               IF (#TMP_dNextTail + 1) >= "DMAXGLASSDATASECTORS" THEN
                   #TMP_dNextTail := 0;
               ELSE
                   #TMP_dNextTail += 1;
               END_IF;

               #TMP_dValue_cmm := #INO_tRibbon.rgtGlassData[#TMP_dSourceIndex].rgtBuffer[#TMP_dNextTail].dEncoderValue_cmm - #INO_tEncoder.dActualEncoderCounter_cmm;

               IF (#TMP_dValue_cmm <= #INO_tRibbon.rgtGlassDataRequest[#TMP_dIndex].IN_dDistanceSnaproll_cmm) THEN

                   #INO_tRibbon.rgtGlassDataRequest[#TMP_dIndex].OUT_dGrossWidth_cmm := #INO_tRibbon.rgtGlassData[#TMP_dSourceIndex].rgtBuffer[#TMP_dNextTail].dGrossWidth_cmm;
                   #INO_tRibbon.rgtGlassDataRequest[#TMP_dIndex].OUT_dNetWidth_cmm := #INO_tRibbon.rgtGlassData[#TMP_dSourceIndex].rgtBuffer[#TMP_dNextTail].dNetWidth_cmm;
                   #INO_tRibbon.rgtGlassDataRequest[#TMP_dIndex].OUT_dGrossWander_cmm := #INO_tRibbon.rgtGlassData[#TMP_dSourceIndex].rgtBuffer[#TMP_dNextTail].dGrossWander_cmm;
                   #INO_tRibbon.rgtGlassDataRequest[#TMP_dIndex].OUT_dNetWander_cmm := #INO_tRibbon.rgtGlassData[#TMP_dSourceIndex].rgtBuffer[#TMP_dNextTail].dNetWander_cmm;

               ELSE
                   EXIT;
               END_IF;

           END_WHILE;
           //Setup data ready
           #INO_tRibbon.rgtGlassDataRequest[#TMP_dIndex].OUT_xDataReady := TRUE;
       END_IF;
   END_FOR;
END_REGION

REGION Network 8 (SCL): Evaluate glass break request
   FOR #TMP_dIndex := 0 TO "DMAXGLASSBREAKREQUEST_IND" DO

       #TMP_xGlassBreak := FALSE;

       IF #INO_tRibbon.rgtGlassBreakRequest[#TMP_dIndex].IN_xRequestGlassBreak AND NOT #INO_tRibbon.rgtGlassBreakRequest[#TMP_dIndex].OUT_xDataReady THEN

           //Evaluate the glass break machine, only the machine before the requested position 
           FOR #TMP_dBreakMachIndex := 0 TO #INO_tRibbon.dActualNumberGlassBreakMachine - 1 DO

               IF (#INO_tRibbon.rgtGlassBreakRequest[#TMP_dIndex].IN_dDistanceSnaproll_cmm >= #INO_tRibbon.rgtGlassBreak[#TMP_dBreakMachIndex].dDistSnapRoll_cmm) THEN
                   CONTINUE;
               END_IF;

               #TMP_xGlassBreak := #INO_tRibbon.rgtGlassBreak[#TMP_dBreakMachIndex].tLastDataBuffer.xGlassBreak;

               #TMP_dNextTail := #INO_tRibbon.rgtGlassBreak[#TMP_dBreakMachIndex].dBufferTail;

               WHILE (#TMP_dNextTail <> #INO_tRibbon.rgtGlassBreak[#TMP_dBreakMachIndex].dBufferHead)
                   AND (#INO_tRibbon.rgtGlassBreak[#TMP_dBreakMachIndex].dBufferHead <> -1) DO

                   IF (#TMP_dNextTail + 1) >= "DMAXGLASSBREAKSECTORS" THEN
                       #TMP_dNextTail := 0;
                   ELSE
                       #TMP_dNextTail += 1;
                   END_IF;

                   #TMP_dValue_cmm := #INO_tRibbon.rgtGlassBreak[#TMP_dBreakMachIndex].rgtBuffer[#TMP_dNextTail].dEncoderValue_cmm - #INO_tEncoder.dActualEncoderCounter_cmm;

                   IF (#TMP_dValue_cmm <= #INO_tRibbon.rgtGlassBreakRequest[#TMP_dIndex].IN_dDistanceSnaproll_cmm) THEN

                       //If the distance is less the snaproll, but greather the safety band. In case of glass break the system will not overwrite the information
                       IF (#TMP_dValue_cmm < #INO_tRibbon.rgtGlassBreakRequest[#TMP_dIndex].IN_dDistanceSnaproll_cmm - #INO_tRibbon.rgtGlassBreakRequest[#TMP_dIndex].IN_dDownstreamOffset_cmm) THEN
                           #TMP_xGlassBreak := #INO_tRibbon.rgtGlassBreak[#TMP_dBreakMachIndex].rgtBuffer[#TMP_dNextTail].xGlassBreak;
                       ELSE
                           IF NOT #TMP_xGlassBreak THEN
                               #TMP_xGlassBreak := #INO_tRibbon.rgtGlassBreak[#TMP_dBreakMachIndex].rgtBuffer[#TMP_dNextTail].xGlassBreak;
                           END_IF;
                       END_IF;

                   ELSE

                       //The position is greather, but still on the position window
                       IF (#TMP_dValue_cmm <= #INO_tRibbon.rgtGlassBreakRequest[#TMP_dIndex].IN_dDistanceSnaproll_cmm + #INO_tRibbon.rgtGlassBreakRequest[#TMP_dIndex].IN_dUpstreamOffset_cmm) THEN
                           IF NOT #TMP_xGlassBreak THEN
                               #TMP_xGlassBreak := #INO_tRibbon.rgtGlassBreak[#TMP_dBreakMachIndex].rgtBuffer[#TMP_dNextTail].xGlassBreak;
                           END_IF;
                       ELSE
                           EXIT; //Exit the while
                       END_IF;

                   END_IF;

               END_WHILE;

               IF #TMP_xGlassBreak THEN
                   EXIT;
               END_IF;
           END_FOR;

           #INO_tRibbon.rgtGlassBreakRequest[#TMP_dIndex].OUT_xDataReady := TRUE;
           #INO_tRibbon.rgtGlassBreakRequest[#TMP_dIndex].OUT_xGlassBreak := #TMP_xGlassBreak;

       END_IF;
   END_FOR;
END_REGION
END_FUNCTION_BLOCK

// folder: 03_Programs_Logics/MCC1200/18_ISRA

FUNCTION_BLOCK "FB_ISRA5D"   // FB21, LAD
{ S7_Optimized_Access := 'TRUE' }
VERSION : 0.1
   VAR_INPUT
      IN_xCycleON : Bool;   // Cycle ON
      IN_xCycleONDel : Bool;   // Delayed cycle ON signal
      IN_dGlassBreakIndexGet : DInt;   // Glass break index get
      IN_xGeneralReset : Bool;   // General reset
      IN_xResetAlarms : Bool;   // Reset alarms
      IN_xFaultsEnabled : Bool;   // Faults enabled
      IN_tInterfaceID : Hw_Any;   // Interface ID
      IN_tID : Conn_Ouc;   // Connection ID
      IN_uiLocalPort : UInt;   // Local port
      IN_dGlassDataMachineIndex : DInt;   // Glass data machine index
      IN_dGlassDataUpdateMachineIndex : DInt;   // Glass data update machine index
      IN_xSimulationActive : Bool;   // Enable simulation (EXPERT USER)
      IN_xScannerON : Bool;
   END_VAR
   VAR_OUTPUT
      OUT_xGlassBreak : Bool;
   END_VAR
   VAR_IN_OUT
      INO_tFBAddDefect : "FB_Defects_Add_V1.00";   // Add defect on buffer
      INO_xDefectBufferFull : Bool;   // Defect buffer full
      INO_tEncoder : "UDT_Encoder";   // Encoder data
      INO_tRibbon : "UDT_RibbonData";   // Ribbon data
      INO_tOptManager : "FB_OptManager_V1.00";   // Optimizer manager
      INO_tCaps : "UDT_CapData_Tracking";   // Caps data
      INO_OB_Init : "GP_OB_Initialize";
   END_VAR
   VAR
      tALM : Struct   // HMI Alarms
         tS : Struct   // Stopping faults
            xNotSyncro : Bool;   // Machine not syncronized {X|X|X|X|O}
            xScannerNotConnected : Bool;   // Scanner not connected {X|X|X|X|O}
            xSpare_2 : Bool;
            xSpare_3 : Bool;
            xSpare_4 : Bool;
            xSpare_5 : Bool;
            xSpare_6 : Bool;
            xSpare_7 : Bool;
            xSpare_8 : Bool;
            xSpare_9 : Bool;
            xSpare_10 : Bool;
            xSpare_11 : Bool;
            xSpare_12 : Bool;
            xSpare_13 : Bool;
            xSpare_14 : Bool;
            xSpare_15 : Bool;
            xSpare_16 : Bool;
            xSpare_17 : Bool;
            xSpare_18 : Bool;
            xSpare_19 : Bool;
            xSpare_20 : Bool;
            xSpare_21 : Bool;
            xSpare_22 : Bool;
            xSpare_23 : Bool;
            xSpare_24 : Bool;
            xSpare_25 : Bool;
            xSpare_26 : Bool;
            xSpare_27 : Bool;
            xSpare_28 : Bool;
            xSpare_29 : Bool;
            xSpare_30 : Bool;
            xSpare_31 : Bool;
         END_STRUCT;
         tF : Struct   // Faults
            xUTelMissing : Bool;   // U telegram missing {X|X|X|X|O}
            xSTelMissing : Bool;   // S telegram missing {X|X|X|X|O}
            xCTelMissing : Bool;   // C telegram missing {X|X|X|X|O}
            xYTelMissing : Bool;   // Y telegram missing {X|X|X|X|O}
            xBTelMissing : Bool;   // B telegram missing {X|X|X|X|O}
            xSpare_5 : Bool;
            xSpare_6 : Bool;
            xSpare_7 : Bool;
            xSpare_8 : Bool;
            xSpare_9 : Bool;
            xSpare_10 : Bool;
            xSpare_11 : Bool;
            xSpare_12 : Bool;
            xSpare_13 : Bool;
            xSpare_14 : Bool;
            xSpare_15 : Bool;
            xSpare_16 : Bool;
            xSpare_17 : Bool;
            xSpare_18 : Bool;
            xSpare_19 : Bool;
            xSpare_20 : Bool;
            xSpare_21 : Bool;
            xSpare_22 : Bool;
            xSpare_23 : Bool;
            xSpare_24 : Bool;
            xSpare_25 : Bool;
            xSpare_26 : Bool;
            xSpare_27 : Bool;
            xSpare_28 : Bool;
            xSpare_29 : Bool;
            xSpare_30 : Bool;
            xSpare_31 : Bool;
         END_STRUCT;
         tW : Struct   // Warnings
            xSpare_0 : Bool;
            xSpare_1 : Bool;
            xSpare_2 : Bool;
            xSpare_3 : Bool;
            xSpare_4 : Bool;
            xSpare_5 : Bool;
            xSpare_6 : Bool;
            xSpare_7 : Bool;
            xSpare_8 : Bool;
            xSpare_9 : Bool;
            xSpare_10 : Bool;
            xSpare_11 : Bool;
            xSpare_12 : Bool;
            xSpare_13 : Bool;
            xSpare_14 : Bool;
            xSpare_15 : Bool;
            xSpare_16 : Bool;
            xSpare_17 : Bool;
            xSpare_18 : Bool;
            xSpare_19 : Bool;
            xSpare_20 : Bool;
            xSpare_21 : Bool;
            xSpare_22 : Bool;
            xSpare_23 : Bool;
            xSpare_24 : Bool;
            xSpare_25 : Bool;
            xSpare_26 : Bool;
            xSpare_27 : Bool;
            xSpare_28 : Bool;
            xSpare_29 : Bool;
            xSpare_30 : Bool;
            xSpare_31 : Bool;
         END_STRUCT;
      END_STRUCT;
   END_VAR
   VAR RETAIN
      tHMR : Struct
         dInspectionStatus : DInt;   // Inspection status (1=Disabled 3=Enabled 4=Wait first syncro 7=Anomaly ) {X|X|X|X|O}
         xScannerON : Bool;   // xScannerON {X|X|X|X|O}
         dDistSnapRoll_cmm : DInt;   // Distance from snaproll [mm/100] {mm/100|mm|X|X|O}
         dDistCenterLine_cmm : DInt;   // Distance from center line [mm/100] {mm/100|mm|X|X|O}
         dCurrentGrossWidth_cmm : DInt;   // Gross width [mm/100] {mm/100|mm|X|X|O}
         dCurrentNetWidth_cmm : DInt;   // Net width [mm/100] {mm/100|mm|X|X|O}
         dCurrentGrossWander_cmm : DInt;   // Gross wander [mm/100] {mm/100|mm|X|X|O}
         dCurrentNetWander_cmm : DInt;   // Net wander [mm/100] {mm/100|mm|X|X|O}
      END_STRUCT;
      tHMW : Struct   // HMI Write
         xAutoInspEnabled : Bool;   // Automatic inspection enabled {X|X|X|X|O}
         xUpdDistSnaproll : Bool;   // Update distance from snaproll {X|X|X|X|O}
         xUpdDistCenterLine : Bool;   // Update distance from center line {X|X|X|X|O}
         xCalibPosition : Bool;   // Calibrate defect position {X|X|X|X|O}
         dCalibDefRealXPos_cmm : DInt;   // Calibration defect real X position [mm/100] {mm/100|mm|0|7000|O}
         dCalibDefRealYPos_cmm : DInt;   // Calibration defect real Y position [mm/100] {mm/100|mm|0|4000|O}
         dCalibDefTeoXPos_cmm : DInt;   // Calibration defect theorical X position [mm/100] {mm/100|mm|0|7000|O}
         dCalibDefTeoYPos_cmm : DInt;   // Calibration defect theorical Y position [mm/100] {mm/100|mm|0|4000|O}
         dDistSnapRoll_cmm : DInt;   // Distance from snaproll [mm/100] {mm/100|mm|0|70000|O}
         dDistCenterLine_cmm : DInt;   // Distance from center line [mm/100] {mm/100|mm|-4000|4000|O}
      END_STRUCT;
   END_VAR
   VAR
      tPhNet : Struct   // Network phases
         xSendInProgress : Bool;   // Send data in progress
         xEndSendInProgress : Bool;   // End send data in progress
         xSpare_2 : Bool;
         xSpare_3 : Bool;
         xSpare_4 : Bool;
         xSpare_5 : Bool;
         xSpare_6 : Bool;
         xSpare_7 : Bool;
         xSpare_8 : Bool;
         xSpare_9 : Bool;
         xSpare_10 : Bool;
         xSpare_11 : Bool;
         xSpare_12 : Bool;
         xSpare_13 : Bool;
         xSpare_14 : Bool;
         xSpare_15 : Bool;
         xSpare_16 : Bool;
         xSpare_17 : Bool;
         xSpare_18 : Bool;
         xSpare_19 : Bool;
         xSpare_20 : Bool;
         xSpare_21 : Bool;
         xSpare_22 : Bool;
         xSpare_23 : Bool;
         xSpare_24 : Bool;
         xSpare_25 : Bool;
         xSpare_26 : Bool;
         xSpare_27 : Bool;
         xSpare_28 : Bool;
         xSpare_29 : Bool;
         xSpare_30 : Bool;
         xSpare_31 : Bool;
      END_STRUCT;
      tPh : Struct   // Machine phases
         xWaitSyncroData : Bool;   // Wait syncro data
         xEndWaitSyncroData : Bool;   // End wait syncro data
         xSpare_2 : Bool;
         xSpare_3 : Bool;
         xSpare_4 : Bool;
         xSpare_5 : Bool;
         xSpare_6 : Bool;
         xSpare_7 : Bool;
         xSpare_8 : Bool;
         xSpare_9 : Bool;
         xSpare_10 : Bool;
         xSpare_11 : Bool;
         xSpare_12 : Bool;
         xSpare_13 : Bool;
         xSpare_14 : Bool;
         xSpare_15 : Bool;
         xSpare_16 : Bool;
         xSpare_17 : Bool;
         xSpare_18 : Bool;
         xSpare_19 : Bool;
         xSpare_20 : Bool;
         xSpare_21 : Bool;
         xSpare_22 : Bool;
         xSpare_23 : Bool;
         xSpare_24 : Bool;
         xSpare_25 : Bool;
         xSpare_26 : Bool;
         xSpare_27 : Bool;
         xSpare_28 : Bool;
         xSpare_29 : Bool;
         xSpare_30 : Bool;
         xSpare_31 : Bool;
      END_STRUCT;
      ST_xMachineSyncronized : Bool;   // Machine is syncronized
      ST_xStoppedFaults : Bool;   // Stopped faults
      ST_xFaults : Bool;   // Faults
      ST_xWarning : Bool;   // Warnings
      ST_xGlassBreak : Bool;   // Glass break
      OS_xSyncroOutLimits : Bool;   // OS.Syncro outside limits
      OS_xSyncroTimeout : Bool;   // OS.Syncro timeout
      AUX_xTelegramError : Bool;   // Telegram error
      AUX_xTelegramYError : Bool;   // Telegram Y error
      AUX_xTelegramBError : Bool;   // Telegram B error
      AUX_xTelegramCError : Bool;   // Telegram C error
      AUX_xTelegramSError : Bool;   // Telegram S error
      AUX_xTelegramUError : Bool;   // Telegram U error
      AUX_xTelegramYMissing : Bool;   // Telegram Y missing
      AUX_xTelegramBMissing : Bool;   // Telegram B missing
      AUX_xTelegramCMissing : Bool;   // Telegram C missing
      AUX_xTelegramSMissing : Bool;   // Telegram S missing
      AUX_xTelegramUMissing : Bool;   // Telegram U missing
      AUX_tUTelegram : Struct   // U telegram
         dTelCounter : DInt;   // Telegram counter [0..65535]
         dFeedPulse_mm : DInt;   // Feeding pulse counter [mm]
         dDefPos_mm : DInt;   // Defect position [mm]
         dDefLengthTot_um : DInt;   // Defect length total [um]
         dDefWidthTot_um : DInt;   // Defect width total [um]
         dDefLengthCore_um : DInt;   // Defect length core [um]
         dDefWidthCore_um : DInt;   // Defect width core [um]
         dDefLengthDef_um : DInt;   // Defect length deformation [um]
         dDefWidthDef_um : DInt;   // Defect width deformation [um]
         dClass : DInt;   // Defect class [01..99]
         dType : DInt;   // Defect type [01..99]
         dPLCPosCount_cmm : DInt;   // PLC Position counter [mm/100]
         dPLCYPos_cmm : DInt;   // PLC Y position value [mm/100]
         strDefectID : String;   // Defect ID string
      END_STRUCT;
      AUX_tYTelegram : Struct   // Y telegram
         dTelCounter : DInt;   // Telegram counter [0..65535]
         dFeedPulse_mm : DInt;   // Feeding pulse counter [mm]
         dInLimit_mm : DInt;   // Inner limit of the observation area [mm]
         dOutLimit_mm : DInt;   // Outer limit o fthe observation area [mm]
         dInLimitUsable_mm : DInt;   // Inner limit of the usable glass width [mm]
         dOutLimitUsable_mm : DInt;   // Outer limit of the usable glass width [mm]
         dInLimitGross_mm : DInt;   // Inner gross glass width [mm]
         dOutLimitGross_mm : DInt;   // Outer gross glass width [mm]
         dCenterOrientInTop_mm : DInt;   // Center orientated position of the inner toproller [mm]
         dEdgeOrientInTop_mm : DInt;   // Edge orientated position of the inner toproller [mm]
         dCenterOrientOutTop_mm : DInt;   // Center orientated position of the outer toproller [mm]
         dEdgeOrientOutTop_mm : DInt;   // Edge orientated position of the outer toproll [mm]
         dPLCPosCount_cmm : DInt;   // PLC Position counter [mm/100]
         dPLCYPos_cmm : DInt;   // PLC Y position value [mm/100]
      END_STRUCT;
      AUX_tCTelegram : Struct   // C Telegram
         dTelCounter : DInt;   // Telegram counter [0..65535]
         dFeedPulseStart_mm : DInt;   // Feeding pulse start counter [mm]
         dFeedPulseEnd_mm : DInt;   // Feeding pulse end counter [mm]
         dBeginAreaY_mm : DInt;   // Begin area Y [mm]
         dEndAreaY_mm : DInt;   // End area Y [mm]
         dPLCPosCountStart_cmm : DInt;   // PLC Position counter start [mm/100]
         dPLCPosCountEnd_cmm : DInt;   // PLC Position counter end [mm/100]
         dPLCYPosStart_cmm : DInt;   // PLC Y position value start [mm/100]
         dPLCYPosEnd_cmm : DInt;   // PLC Y position value end [mm/100]
         dPLCClusterLength_um : DInt;   // PLC Cluster length [um]
         dPLCClusterWidth_um : DInt;   // PLC Cluster width [um]
      END_STRUCT;
      AUX_tBTelegram : Struct   // B Telegram
         dTelCounter : DInt;   // Telegram counter [0..65535]
         dFeedPulse_mm : DInt;   // Feeding pulse counter [mm]
         xNewTelegram : Bool;   // New telegram received
      END_STRUCT;
      AUX_tSTelegram : Struct   // S Telegram
         dTelCounter : DInt;   // Telegram counter [0..65535]
         dFeedPulse_mm : DInt;   // Feeding pulse counter [mm]
         xNewTelegram : Bool;   // New telegram received
      END_STRUCT;
      AUX_tWTelegram : Struct   // T Telegram
         dTelCounter : DInt;   // Telegram counter [0..65535]
         dFeedPulse_mm : DInt;   // Feeding pulse counter [mm]
         dGrossWidthMin_mm : DInt;   // Gross width min [mm]
         dGrossWidthMax_mm : DInt;   // Gross width max [mm]
         dCutToolOpSide_mm : DInt;   // Cut tool opside [mm]
         dCutToolOppoOpSide_mm : DInt;   // Cut tool opposite operator side [mm]
         xNewTelegram : Bool;   // New telegram received
      END_STRUCT;
      AUX_dISRAValidCountMeter_mm : DInt;   // Last valid isra counter on meter [mm]
      AUX_dPLCValidCountMeter_cmm : DInt;   // Last valid PLC counter on meter [mm/100]
      AUX_rgcReceiveBuffer : Array[0..#DRECV_BUFFER_MAX_IND] of Char;   // Receive buffer
      AUX_dNumCharRecvBuffer : DInt;   // Number of char on the receive buffer
      AUX_rgsWTelegram : Array[0..#DNUMCHAR_TEL_W_INDEX] of Char;   // T Telegram char array
      AUX_tConnData : TCON_IP_v4;   // Connection data structure
      FB_TSend : TSEND_C;   // FB send
      FB_TRecv : TRCV_C;   // FB receive
      AUX_xResetSendConnection : Bool;   // Reset send connection
      AUX_rgcReceiveTempBuffer : Array[0..#DRECV_BUFFER_TEMP_IND] of Char;   // Temporary receive buffer
      tmON_SendTimeout : "UDT_IECTON_V1.00";   // Send timeout
      AUX_xSimDecModeGWidth : Bool;   // SIMULATION - Decrement mode gross width
      AUX_xSimIncModeGWidth : Bool;   // SIMULATION - Increment mode gross width
      AUX_xSimDecModeNWidth : Bool;   // SIMULATION - Decrement mode net width
      AUX_xSimIncModeNWidth : Bool;   // SIMULATION - Decrement mode net width
      AUX_xSimDecModeWander : Bool;   // SIMULATION - Decrement mode wander
      AUX_xSimIncModeWander : Bool;   // SIMULATION - Decrement mode wander
   END_VAR
   VAR RETAIN
      AUX_dSimGrossWidth_cmm : DInt;   // SIMULATION - Gross width [mm/100]
      AUX_dSimNetWidth_cmm : DInt;   // SIMULATION - Net width [mm/100]
      AUX_dSimWander_cmm : DInt;   // SIMULATION - Wander [mm/100]
   END_VAR
   VAR_TEMP
      TMP_dwValue : DWord;
      TMP_dIndex : DInt;
      TMP_dCharCounter : DInt;
      TMP_dTelCount : DInt;
      TMP_strValue : String;
      TMP_dCountPos_cmm : DInt;
      TMP_iRetVal : Int;
      TMP_dValue_cmm : DInt;
      TMP_xDummy : Bool;
      TMP_iStrLength : Int;
      TMP_uiMovedChar : UInt;
      TMP_xEnableReceive : Bool;
   END_VAR
   VAR CONSTANT
      DRECV_BUFFER_MAX : DInt := 5000;   // Maximum number of character on the receive buffer
      DRECV_BUFFER_MAX_IND : DInt := 4999;   // Maximum number of character on the receive buffer index
      DRECV_BUFFER_TEMP : DInt := 1000;   // Maximum number of character on the temporary receive buffer
      DRECV_BUFFER_TEMP_IND : DInt := 999;   // Maximum number of character on the temporary receive buffer index
      STR_CR : Char := '$R';   // CR
      STR_LF : Char := '$L';   // LF
      DNUMCHAR_TEL_U : DInt := 106;   // Number of char U telegram
      DNUMCHAR_TEL_C : DInt := 36;   // Number of char C telegram
      DNUMCHAR_TEL_Y : DInt := 75;   // Number of char Y telegram
      DNUMCHAR_TEL_B_S : DInt := 15;   // Number of char B - S telegram
      DCLUSTER_CLASS : DInt := 21;   // Cluster defect used class
      DCLUSTER_SUBTYPE : DInt := 1004;   // Cluster defect subtype
      DNUMCHAR_TEL_W : DInt := 39;   // Number of char W telegram
      DNUMCHAR_TEL_W_INDEX : DInt := 38;   // Number of char W telegram index
      DISRADEADPOINT_CMM : DInt := 250000;   // ISRA Dead point position quota [mm/100]
      CONST_DBREAKDOWNOFF_CMM : DInt := 100000;   // Break downstream offset [mm/100]
      CONST_DBREAKUPOFF_CMM : DInt := 100000;   // Break upstream offset [mm/100]
      BCONNTYPE : Byte := 16#0B;   // Optimizer connection type
      DSIM_MINGROSSWIDTH_CMM : DInt := 340000;   // Simulation minimum gross width [mm/100]
      DSIM_MAXGROSSWIDTH_CMM : DInt := 350000;   // Simulation maximum gross width [mm/100]
      DSIM_MINNETWIDTH_CMM : DInt := 330000;   // Simulation minimum net width [mm/100]
      DSIM_MAXNETWIDTH_CMM : DInt := 340000;   // Simulation maximum net width [mm/100]
      DSIM_MINNETWANDER_CMM : DInt := -20000;   // Simulation minimum net wander [mm/100]
      DSIM_MAXNETWANDER_CMM : DInt := 20000;   // Simulation maximum net wander [mm/100]
   END_VAR
   VAR_TEMP   // added for the SCL form of the ladder/FBD networks
      _w1 : Bool;
   END_VAR
BEGIN

REGION Network 1: ####_CONSTANTS_####
END_REGION

REGION Network 2 (SCL): General reset actions
   IF #IN_xGeneralReset THEN

       #AUX_tConnData.InterfaceId := #IN_tInterfaceID;
       #AUX_tConnData.ID := #IN_tID;
       #AUX_tConnData.ConnectionType := #BCONNTYPE;
       #AUX_tConnData.ActiveEstablished := FALSE;
       #AUX_tConnData.RemotePort := 0;
       #AUX_tConnData.LocalPort := #IN_uiLocalPort;

       #tPh.xWaitSyncroData := FALSE;
       #tPh.xEndWaitSyncroData := FALSE;

       #tPhNet.xSendInProgress := FALSE;
       #tPhNet.xEndSendInProgress := FALSE;

   END_IF;
END_REGION

REGION Network 3: ### ETHERNET RECEIVE DATA ###
END_REGION

REGION Network 4 (SCL): Manage send and receive
   #AUX_xResetSendConnection := #IN_xGeneralReset OR (#FB_TSend.s_TDIAG_Status.State <> b#16#04 AND #IN_xResetAlarms);

   #FB_TSend(REQ:=#tPhNet.xSendInProgress,
             CONT:=TRUE,
             LEN:=0,
             CONNECT:=#AUX_tConnData,
             DATA:=#AUX_rgsWTelegram,
             COM_RST:=#AUX_xResetSendConnection);

   IF (#DRECV_BUFFER_MAX - #AUX_dNumCharRecvBuffer) > #DRECV_BUFFER_TEMP THEN
       #TMP_xEnableReceive := TRUE;
   ELSE
       #TMP_xEnableReceive := FALSE;
   END_IF;

   #FB_TRecv(EN_R:=#TMP_xEnableReceive,
               CONT:=TRUE,
               LEN:=0,
               ADHOC:=TRUE,
               CONNECT:=#AUX_tConnData,
               DATA:=#AUX_rgcReceiveTempBuffer,
               COM_RST:=#AUX_xResetSendConnection);

   IF #FB_TRecv.DONE THEN

       //Copy the received data
       #TMP_iRetVal := MOVE_BLK_VARIANT(SRC:=#AUX_rgcReceiveTempBuffer, COUNT:=#FB_TRecv.RCVD_LEN, SRC_INDEX:=0, DEST_INDEX:=#AUX_dNumCharRecvBuffer, DEST=>#AUX_rgcReceiveBuffer);
       #AUX_dNumCharRecvBuffer += UDINT_TO_DINT(#FB_TRecv.RCVD_LEN);

   END_IF;
END_REGION

REGION Network 5: ####_MATCH_####
END_REGION

REGION Network 6: ####_HMI_LOGICS_####
END_REGION

REGION Network 7 (SCL): Manage HMI
   IF #tHMW.xUpdDistSnaproll THEN
       #tHMW.xUpdDistSnaproll := FALSE;
       #tHMR.dDistSnapRoll_cmm := #tHMW.dDistSnapRoll_cmm;
   END_IF;

   IF #tHMW.xUpdDistCenterLine THEN
       #tHMW.xUpdDistCenterLine := FALSE;
       #tHMR.dDistCenterLine_cmm := #tHMW.dDistCenterLine_cmm;
   END_IF;

   IF #tHMW.xCalibPosition THEN

       IF #tHMR.dDistCenterLine_cmm <= 0 THEN
           #tHMR.dDistCenterLine_cmm := #tHMR.dDistCenterLine_cmm - (#tHMW.dCalibDefTeoYPos_cmm - #tHMW.dCalibDefRealYPos_cmm); 
       ELSE
           #tHMR.dDistCenterLine_cmm := #tHMR.dDistCenterLine_cmm + (#tHMW.dCalibDefRealYPos_cmm - #tHMW.dCalibDefTeoYPos_cmm); 
       END_IF;        

       #tHMR.dDistSnapRoll_cmm := #tHMR.dDistSnapRoll_cmm + (#tHMW.dCalibDefRealXPos_cmm - #tHMW.dCalibDefTeoXPos_cmm);

       #tHMW.dCalibDefRealXPos_cmm := #tHMW.dCalibDefTeoXPos_cmm;
       #tHMW.dCalibDefRealYPos_cmm := #tHMW.dCalibDefTeoYPos_cmm;
       #tHMW.xCalibPosition := FALSE;

   END_IF;

   (*IF #tHMW.xEnAutoInsp THEN
       #tHMW.xEnAutoInsp := FALSE;
       #tHMR.xAutoInspEnabled := TRUE;
   END_IF;

   IF #tHMW.xDisAutoInsp THEN
       #tHMW.xDisAutoInsp := FALSE;
       #tHMR.xAutoInspEnabled := FALSE;
   END_IF; *)
END_REGION

REGION Network 8: ####_ALARMS_####
END_REGION

REGION Network 9 (SCL): Reset alarms
   IF #IN_xResetAlarms THEN

       #TMP_dwValue := 0;

       SCATTER(IN:=#TMP_dwValue,
               OUT=>#tALM.tS);

       SCATTER(IN:=#TMP_dwValue,
               OUT=>#tALM.tF);

       SCATTER(IN:=#TMP_dwValue,
               OUT=>#tALM.tW);


   END_IF;
END_REGION

REGION Network 10: Machine not syncronized {X|X|X|X|O}
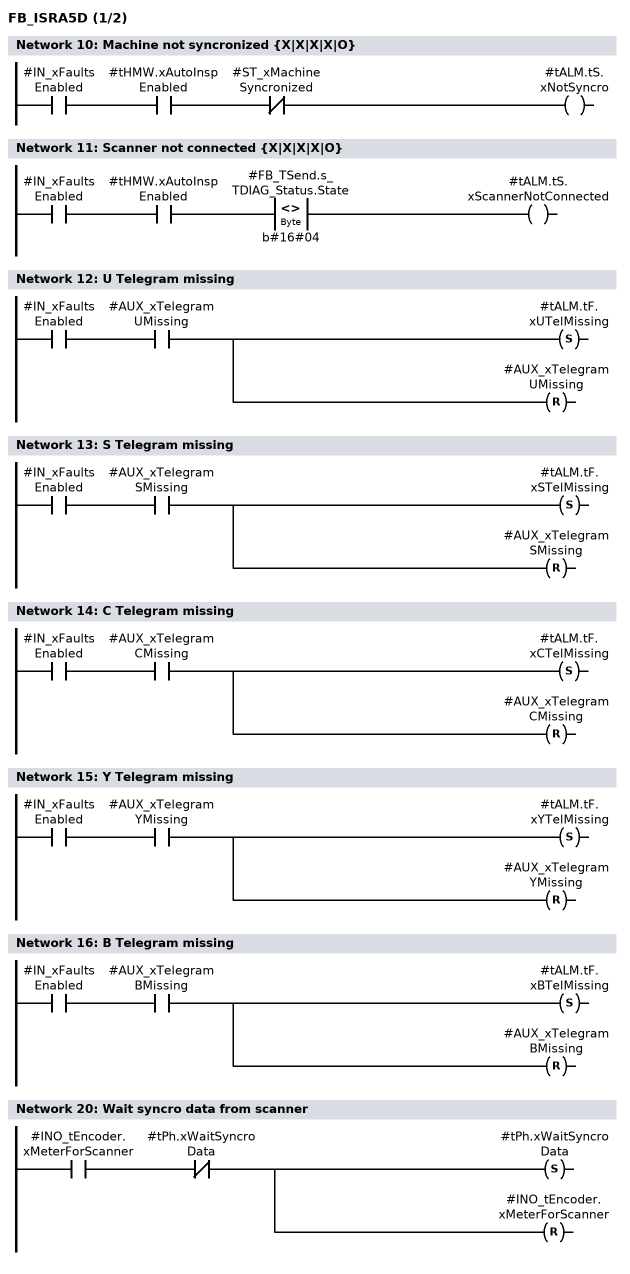
   RUNG wire#powerrail
      Contact( #IN_xFaultsEnabled )
      Contact( #tHMW.xAutoInspEnabled )
      I_Contact( #ST_xMachineSyncronized )
      Coil( #tALM.tS.xNotSyncro )
   END_RUNG
   // the same network as SCL:
   #tALM.tS.xNotSyncro := #IN_xFaultsEnabled AND #tHMW.xAutoInspEnabled AND NOT #ST_xMachineSyncronized;
END_REGION

REGION Network 11: Scanner not connected {X|X|X|X|O}
   RUNG wire#powerrail
      Contact( #IN_xFaultsEnabled )
      Contact( #tHMW.xAutoInspEnabled )
      { S7_Templates := "SrcType := Byte" } NE_Contact(in1 := #FB_TSend.s_TDIAG_Status.State, in2 := b#16#04)
      Coil( #tALM.tS.xScannerNotConnected )
   END_RUNG
   // the same network as SCL:
   #tALM.tS.xScannerNotConnected := #IN_xFaultsEnabled AND #tHMW.xAutoInspEnabled AND (#FB_TSend.s_TDIAG_Status.State <> b#16#04);
END_REGION

REGION Network 12: U Telegram missing
   RUNG wire#powerrail
      Contact( #IN_xFaultsEnabled )
      Contact( #AUX_xTelegramUMissing )
      wire#w1
      S_Coil( #tALM.tF.xUTelMissing )
   END_RUNG
   RUNG wire#w1
      R_Coil( #AUX_xTelegramUMissing )
   END_RUNG
   // the same network as SCL:
   IF #IN_xFaultsEnabled AND #AUX_xTelegramUMissing THEN
       #tALM.tF.xUTelMissing := TRUE;
       #AUX_xTelegramUMissing := FALSE;
   END_IF;
END_REGION

REGION Network 13: S Telegram missing
   RUNG wire#powerrail
      Contact( #IN_xFaultsEnabled )
      Contact( #AUX_xTelegramSMissing )
      wire#w1
      S_Coil( #tALM.tF.xSTelMissing )
   END_RUNG
   RUNG wire#w1
      R_Coil( #AUX_xTelegramSMissing )
   END_RUNG
   // the same network as SCL:
   IF #IN_xFaultsEnabled AND #AUX_xTelegramSMissing THEN
       #tALM.tF.xSTelMissing := TRUE;
       #AUX_xTelegramSMissing := FALSE;
   END_IF;
END_REGION

REGION Network 14: C Telegram missing
   RUNG wire#powerrail
      Contact( #IN_xFaultsEnabled )
      Contact( #AUX_xTelegramCMissing )
      wire#w1
      S_Coil( #tALM.tF.xCTelMissing )
   END_RUNG
   RUNG wire#w1
      R_Coil( #AUX_xTelegramCMissing )
   END_RUNG
   // the same network as SCL:
   IF #IN_xFaultsEnabled AND #AUX_xTelegramCMissing THEN
       #tALM.tF.xCTelMissing := TRUE;
       #AUX_xTelegramCMissing := FALSE;
   END_IF;
END_REGION

REGION Network 15: Y Telegram missing
   RUNG wire#powerrail
      Contact( #IN_xFaultsEnabled )
      Contact( #AUX_xTelegramYMissing )
      wire#w1
      S_Coil( #tALM.tF.xYTelMissing )
   END_RUNG
   RUNG wire#w1
      R_Coil( #AUX_xTelegramYMissing )
   END_RUNG
   // the same network as SCL:
   IF #IN_xFaultsEnabled AND #AUX_xTelegramYMissing THEN
       #tALM.tF.xYTelMissing := TRUE;
       #AUX_xTelegramYMissing := FALSE;
   END_IF;
END_REGION

REGION Network 16: B Telegram missing
   RUNG wire#powerrail
      Contact( #IN_xFaultsEnabled )
      Contact( #AUX_xTelegramBMissing )
      wire#w1
      S_Coil( #tALM.tF.xBTelMissing )
   END_RUNG
   RUNG wire#w1
      R_Coil( #AUX_xTelegramBMissing )
   END_RUNG
   // the same network as SCL:
   IF #IN_xFaultsEnabled AND #AUX_xTelegramBMissing THEN
       #tALM.tF.xBTelMissing := TRUE;
       #AUX_xTelegramBMissing := FALSE;
   END_IF;
END_REGION

REGION Network 17 (SCL): Calculate comulative statuses
       GATHER(IN:=#tALM.tS,
              OUT=>#TMP_dwValue);

       IF #TMP_dwValue <> 0 THEN
           #ST_xStoppedFaults := TRUE;
       ELSE
           #ST_xStoppedFaults := FALSE;
       END_IF;

       GATHER(IN:=#tALM.tF,
              OUT=>#TMP_dwValue);

       IF #TMP_dwValue <> 0 THEN
           #ST_xFaults := TRUE;
       ELSE
           #ST_xFaults := FALSE;
       END_IF;

       GATHER(IN:=#tALM.tW,
              OUT=>#TMP_dwValue);

       IF #TMP_dwValue <> 0 THEN
           #ST_xWarning := TRUE;
       ELSE
           #ST_xWarning := FALSE;
       END_IF;
END_REGION

REGION Network 18: ### PHASES AND LOGICS ###
END_REGION

REGION Network 19 (SCL): Search packet
   #TMP_dCharCounter := 1;
   #TMP_dIndex := 0;
   WHILE (#TMP_dIndex <= #AUX_dNumCharRecvBuffer - 2)  DO

       #TMP_dCharCounter += 1;

       //Loop until to find one CR + LF
       IF #AUX_rgcReceiveBuffer[#TMP_dIndex] = #STR_CR AND #AUX_rgcReceiveBuffer[#TMP_dIndex + 1] = #STR_LF THEN

           CASE #TMP_dCharCounter OF
             #DNUMCHAR_TEL_U:

               IF  #AUX_rgcReceiveBuffer[0] = 'U' AND
                   #AUX_rgcReceiveBuffer[1] = ' ' AND
                   #AUX_rgcReceiveBuffer[7] = ' ' AND
                   #AUX_rgcReceiveBuffer[13] = ' ' AND
                   #AUX_rgcReceiveBuffer[19] = ' ' AND
                   #AUX_rgcReceiveBuffer[27] = ' ' AND
                   #AUX_rgcReceiveBuffer[35] = ' ' AND
                   #AUX_rgcReceiveBuffer[43] = ' ' AND
                   #AUX_rgcReceiveBuffer[51] = ' ' AND
                   #AUX_rgcReceiveBuffer[59] = ' ' AND
                   #AUX_rgcReceiveBuffer[67] = ' ' AND
                   #AUX_rgcReceiveBuffer[70] = ' ' AND
                   #AUX_rgcReceiveBuffer[73] = ' ' AND
                   #AUX_rgcReceiveBuffer[104] = #STR_CR AND
                   #AUX_rgcReceiveBuffer[105] = #STR_LF THEN

                   //Evaluate the data of the U telegram
                   #TMP_dTelCount :=  #AUX_tUTelegram.dTelCounter;               

                   #TMP_dTelCount += 1;

                   IF #TMP_dTelCount >= 65535 THEN
                       #TMP_dTelCount := 1;
                   END_IF; 

                   Chars_TO_Strg(Chars:=#AUX_rgcReceiveBuffer,
                                 pChars:=2,
                                 Cnt:=5,
                                 Strg=>#TMP_strValue);

                   #AUX_tUTelegram.dTelCounter := STRING_TO_DINT(#TMP_strValue); 

                   IF (#TMP_dTelCount <> #AUX_tUTelegram.dTelCounter) THEN
                       #AUX_xTelegramUMissing := 1;    
                   END_IF;

                   //Feeding pulse counter
                   Chars_TO_Strg(Chars:=#AUX_rgcReceiveBuffer,
                                 pChars:=8,
                                 Cnt:=5,
                                 Strg=>#TMP_strValue);

                   #AUX_tUTelegram.dFeedPulse_mm := STRING_TO_DINT(#TMP_strValue); 

                   //Defect position
                   Chars_TO_Strg(Chars:=#AUX_rgcReceiveBuffer,
                                 pChars:=14,
                                 Cnt:=5,
                                 Strg=>#TMP_strValue);

                   #AUX_tUTelegram.dDefPos_mm := STRING_TO_DINT(#TMP_strValue); 

                   //Defect length total
                   Chars_TO_Strg(Chars:=#AUX_rgcReceiveBuffer,
                                 pChars:=20,
                                 Cnt:=7,
                                 Strg=>#TMP_strValue);

                   #AUX_tUTelegram.dDefLengthTot_um := STRING_TO_DINT(#TMP_strValue); 

                   //Defect width total
                   Chars_TO_Strg(Chars:=#AUX_rgcReceiveBuffer,
                                 pChars:=28,
                                 Cnt:=7,
                                 Strg=>#TMP_strValue);

                   #AUX_tUTelegram.dDefWidthTot_um := STRING_TO_DINT(#TMP_strValue); 

                   //Defect length core
                   Chars_TO_Strg(Chars:=#AUX_rgcReceiveBuffer,
                                 pChars:=36,
                                 Cnt:=7,
                                 Strg=>#TMP_strValue);

                   #AUX_tUTelegram.dDefLengthCore_um := STRING_TO_DINT(#TMP_strValue); 

                   //Defect width core
                   Chars_TO_Strg(Chars:=#AUX_rgcReceiveBuffer,
                                 pChars:=44,
                                 Cnt:=7,
                                 Strg=>#TMP_strValue);

                   #AUX_tUTelegram.dDefWidthCore_um := STRING_TO_DINT(#TMP_strValue); 

                   //Defect length deformation
                   Chars_TO_Strg(Chars:=#AUX_rgcReceiveBuffer,
                                 pChars:=52,
                                 Cnt:=7,
                                 Strg=>#TMP_strValue);

                   #AUX_tUTelegram.dDefLengthDef_um := STRING_TO_DINT(#TMP_strValue); 

                   //Defect width deformation
                   Chars_TO_Strg(Chars:=#AUX_rgcReceiveBuffer,
                                 pChars:=60,
                                 Cnt:=7,
                                 Strg=>#TMP_strValue);

                   #AUX_tUTelegram.dDefWidthDef_um := STRING_TO_DINT(#TMP_strValue); 

                   //Defect class
                   Chars_TO_Strg(Chars:=#AUX_rgcReceiveBuffer,
                                 pChars:=68,
                                 Cnt:=2,
                                 Strg=>#TMP_strValue);

                   #AUX_tUTelegram.dClass := STRING_TO_DINT(#TMP_strValue); 

                   //Defect type
                   Chars_TO_Strg(Chars:=#AUX_rgcReceiveBuffer,
                                 pChars:=71,
                                 Cnt:=2,
                                 Strg=>#TMP_strValue);

                   //Defect ID 
                   Chars_TO_Strg(Chars:=#AUX_rgcReceiveBuffer,
                                 pChars:=74,
                                 Cnt:=30,
                                 Strg=>#AUX_tUTelegram.strDefectID);

                   #AUX_tUTelegram.dType := STRING_TO_DINT(#TMP_strValue); 

                   //Check the conformity
                   IF #AUX_tUTelegram.dTelCounter < 0 OR 
                      #AUX_tUTelegram.dTelCounter > 65535 OR
                      #AUX_tUTelegram.dFeedPulse_mm < 0 OR 
                      #AUX_tUTelegram.dFeedPulse_mm > 65535 OR
                      #AUX_tUTelegram.dDefPos_mm < 0 OR 
                      #AUX_tUTelegram.dDefPos_mm > 65535 OR
                      #AUX_tUTelegram.dDefLengthTot_um < 0 OR
                      #AUX_tUTelegram.dDefLengthTot_um > 9999999 OR
                      #AUX_tUTelegram.dDefWidthTot_um < 0 OR
                      #AUX_tUTelegram.dDefWidthTot_um > 9999999 OR
                      #AUX_tUTelegram.dDefLengthCore_um < 0 OR
                      #AUX_tUTelegram.dDefLengthCore_um > 9999999 OR
                      #AUX_tUTelegram.dDefWidthCore_um < 0 OR
                      #AUX_tUTelegram.dDefWidthCore_um > 9999999 OR 
                      #AUX_tUTelegram.dDefLengthDef_um < 0 OR
                      #AUX_tUTelegram.dDefLengthDef_um > 9999999 OR
                      #AUX_tUTelegram.dDefWidthDef_um < 0 OR
                      #AUX_tUTelegram.dDefWidthDef_um > 9999999 OR
                      #AUX_tUTelegram.dClass < 1 OR
                      #AUX_tUTelegram.dClass > 99 OR
                      #AUX_tUTelegram.dType < 1 OR
                      #AUX_tUTelegram.dType > 99 THEN

                      #AUX_xTelegramUError := TRUE;
                   ELSE

                       IF #ST_xMachineSyncronized AND #tHMW.xAutoInspEnabled THEN
                           #TMP_dCountPos_cmm := #AUX_tUTelegram.dFeedPulse_mm - #AUX_dISRAValidCountMeter_mm;

                           IF #TMP_dCountPos_cmm < -32767 THEN
                               #AUX_tUTelegram.dPLCPosCount_cmm  := #AUX_dPLCValidCountMeter_cmm + ((#TMP_dCountPos_cmm + 65536)*100);
                           ELSIF #TMP_dCountPos_cmm > 32767 THEN
                               #AUX_tUTelegram.dPLCPosCount_cmm  := #AUX_dPLCValidCountMeter_cmm + ((#TMP_dCountPos_cmm - 65536)*100);
                           ELSE
                               #AUX_tUTelegram.dPLCPosCount_cmm := #AUX_dPLCValidCountMeter_cmm + (#TMP_dCountPos_cmm*100);
                           END_IF;

                           IF #tHMR.dDistCenterLine_cmm <= 0 THEN
                               #AUX_tUTelegram.dPLCYPos_cmm := #tHMR.dDistCenterLine_cmm + (#AUX_tUTelegram.dDefPos_mm * 100);      
                           ELSE
                               #AUX_tUTelegram.dPLCYPos_cmm := #tHMR.dDistCenterLine_cmm - (#AUX_tUTelegram.dDefPos_mm * 100);      
                           END_IF;

                           #AUX_tUTelegram.dPLCPosCount_cmm := #tHMR.dDistSnapRoll_cmm + #AUX_tUTelegram.dPLCPosCount_cmm;

                           #INO_tFBAddDefect(IN_dClass:=#AUX_tUTelegram.dClass,
                              IN_dSubType:=#AUX_tUTelegram.dType,
                              IN_dXPosition_cmm:=#AUX_tUTelegram.dPLCPosCount_cmm - (#AUX_tUTelegram.dDefLengthTot_um / 20),
                              IN_dYPosition_cmm:=#AUX_tUTelegram.dPLCYPos_cmm - (#AUX_tUTelegram.dDefWidthTot_um / 20),
                              IN_dTotalLength_um:=#AUX_tUTelegram.dDefLengthTot_um,
                              IN_dTotalWidth_um:=#AUX_tUTelegram.dDefWidthTot_um,
                              IN_dCoreLength_um := #AUX_tUTelegram.dDefLengthCore_um,
                              IN_dCoreWidth_um:=#AUX_tUTelegram.dDefWidthCore_um,
                              IN_dDistLength_um := #AUX_tUTelegram.dDefLengthDef_um,
                              IN_dDistWidth_um:=#AUX_tUTelegram.dDefWidthDef_um,
                              IN_dOptValue_mdptr:=0,
                              OUT_xBufferFull => #INO_xDefectBufferFull,
                              IN_strDefectID:=#AUX_tUTelegram.strDefectID);

                       END_IF;                        

                   END_IF;
               ELSE
                   #AUX_xTelegramUError := TRUE;                    
               END_IF;

             #DNUMCHAR_TEL_C:  

               IF  #AUX_rgcReceiveBuffer[0] = 'C' AND
                   #AUX_rgcReceiveBuffer[1] = ' ' AND
                   #AUX_rgcReceiveBuffer[7] = ' ' AND
                   #AUX_rgcReceiveBuffer[13] = ' ' AND
                   #AUX_rgcReceiveBuffer[19] = ' ' AND
                   #AUX_rgcReceiveBuffer[25] = ' ' AND
                   #AUX_rgcReceiveBuffer[31] = ' ' AND
                   #AUX_rgcReceiveBuffer[34] = #STR_CR AND
                   #AUX_rgcReceiveBuffer[35] = #STR_LF THEN


                   //Evaluate the data of the U telegram
                   #TMP_dTelCount :=  #AUX_tCTelegram.dTelCounter;               

                   #TMP_dTelCount += 1;

                   IF #TMP_dTelCount >= 65535 THEN
                       #TMP_dTelCount := 1;
                   END_IF; 

                   Chars_TO_Strg(Chars:=#AUX_rgcReceiveBuffer,
                                 pChars:=2,
                                 Cnt:=5,
                                 Strg=>#TMP_strValue);

                   #AUX_tCTelegram.dTelCounter := STRING_TO_DINT(#TMP_strValue); 

                   IF (#TMP_dTelCount <> #AUX_tCTelegram.dTelCounter) THEN
                       #AUX_xTelegramCMissing := 1;    
                   END_IF;

                   //Feeding pulse start counter
                   Chars_TO_Strg(Chars:=#AUX_rgcReceiveBuffer,
                                 pChars:=8,
                                 Cnt:=5,
                                 Strg=>#TMP_strValue);

                   #AUX_tCTelegram.dFeedPulseStart_mm := STRING_TO_DINT(#TMP_strValue);

                   //Feeding pulse end counter
                   Chars_TO_Strg(Chars:=#AUX_rgcReceiveBuffer,
                                 pChars:=14,
                                 Cnt:=5,
                                 Strg=>#TMP_strValue);

                   #AUX_tCTelegram.dFeedPulseEnd_mm := STRING_TO_DINT(#TMP_strValue);

                   //Begin area Y 
                   Chars_TO_Strg(Chars:=#AUX_rgcReceiveBuffer,
                                 pChars:=20,
                                 Cnt:=5,
                                 Strg=>#TMP_strValue);

                   #AUX_tCTelegram.dBeginAreaY_mm := STRING_TO_DINT(#TMP_strValue);

                   //End area Y 
                   Chars_TO_Strg(Chars:=#AUX_rgcReceiveBuffer,
                                 pChars:=26,
                                 Cnt:=5,
                                 Strg=>#TMP_strValue);

                   #AUX_tCTelegram.dEndAreaY_mm := STRING_TO_DINT(#TMP_strValue);

                   //Check the conformity
                   IF  #AUX_tCTelegram.dTelCounter < 0 OR 
                       #AUX_tCTelegram.dTelCounter > 65535 OR
                       #AUX_tCTelegram.dFeedPulseStart_mm < 0 OR 
                       #AUX_tCTelegram.dFeedPulseStart_mm > 65535 OR 
                       #AUX_tCTelegram.dFeedPulseEnd_mm < 0 OR 
                       #AUX_tCTelegram.dFeedPulseEnd_mm > 65535 OR
                       #AUX_tCTelegram.dBeginAreaY_mm < 0 OR 
                       #AUX_tCTelegram.dBeginAreaY_mm > 9999999 OR
                       #AUX_tCTelegram.dEndAreaY_mm < 0 OR 
                       #AUX_tCTelegram.dEndAreaY_mm > 9999999 THEN

                       #AUX_xTelegramCError := 1;  

                   ELSE
                       IF #ST_xMachineSyncronized AND #tHMW.xAutoInspEnabled THEN

                           #TMP_dCountPos_cmm := #AUX_tCTelegram.dFeedPulseStart_mm - #AUX_dISRAValidCountMeter_mm;

                           IF #TMP_dCountPos_cmm < -32767 THEN
                               #AUX_tCTelegram.dPLCPosCountStart_cmm  := #AUX_dPLCValidCountMeter_cmm + (#TMP_dCountPos_cmm + 65536);
                           ELSIF #TMP_dCountPos_cmm > 32767 THEN
                               #AUX_tCTelegram.dPLCPosCountStart_cmm  := #AUX_dPLCValidCountMeter_cmm + (#TMP_dCountPos_cmm - 65536);
                           ELSE
                               #AUX_tCTelegram.dPLCPosCountStart_cmm := #AUX_dPLCValidCountMeter_cmm + #TMP_dCountPos_cmm;
                           END_IF;

                           IF #tHMR.dDistCenterLine_cmm <= 0 THEN
                               #AUX_tCTelegram.dPLCYPosStart_cmm := #tHMR.dDistCenterLine_cmm + (#AUX_tCTelegram.dBeginAreaY_mm * 100);     
                               #AUX_tCTelegram.dPLCYPosEnd_cmm := #tHMR.dDistCenterLine_cmm + (#AUX_tCTelegram.dEndAreaY_mm * 100);     
                           ELSE
                               #AUX_tCTelegram.dPLCYPosStart_cmm := #tHMR.dDistCenterLine_cmm - (#AUX_tCTelegram.dEndAreaY_mm * 100);       
                               #AUX_tCTelegram.dPLCYPosStart_cmm := #tHMR.dDistCenterLine_cmm - (#AUX_tCTelegram.dBeginAreaY_mm * 100);     
                           END_IF;

                           #AUX_tCTelegram.dPLCPosCountStart_cmm := #tHMR.dDistSnapRoll_cmm + #AUX_tCTelegram.dPLCPosCountStart_cmm;
                           #AUX_tCTelegram.dPLCPosCountEnd_cmm := #tHMR.dDistSnapRoll_cmm + #AUX_tCTelegram.dPLCPosCountEnd_cmm;
                           #AUX_tCTelegram.dPLCClusterLength_um := (#AUX_tCTelegram.dPLCPosCountEnd_cmm -  #AUX_tCTelegram.dPLCPosCountStart_cmm) * 10;
                           #AUX_tCTelegram.dPLCClusterWidth_um := (#AUX_tCTelegram.dPLCYPosEnd_cmm - #AUX_tCTelegram.dPLCYPosStart_cmm) * 10;

                         //  #INO_tFBAddDefect(IN_dClass:=#DCLUSTER_CLASS,
                         //     IN_dSubType:=#DCLUSTER_SUBTYPE,
                         //     IN_dXPosition_cmm:=#AUX_tCTelegram.dPLCPosCountStart_cmm,
                         //     IN_dYPosition_cmm:=#AUX_tCTelegram.dPLCYPosStart_cmm,
                         //     IN_dTotalLength_um:=#AUX_tCTelegram.dPLCClusterLength_um,
                         //     IN_dTotalWidth_um:=#AUX_tCTelegram.dPLCClusterWidth_um,
                         //     IN_dCoreLength_um := #AUX_tCTelegram.dPLCClusterLength_um,
                         //     IN_dCoreWidth_um:=#AUX_tCTelegram.dPLCClusterWidth_um,
                         //     IN_dDistLength_um := #AUX_tCTelegram.dPLCClusterLength_um,
                         //     IN_dDistWidth_um:=#AUX_tCTelegram.dPLCClusterWidth_um,
                         //     IN_dOptValue_mdptr:=0,
                         //     OUT_xBufferFull => #INO_xDefectBufferFull,
                         //     IN_strDefectID:='CLUSTER_DEFECT');

                       END_IF;

                   END_IF;

               ELSE
                   #AUX_xTelegramCError := TRUE;
               END_IF;

             #DNUMCHAR_TEL_Y:

               IF  #AUX_rgcReceiveBuffer[0] = 'Y' AND
                   #AUX_rgcReceiveBuffer[1] = ' ' AND
                   #AUX_rgcReceiveBuffer[7] = ' ' AND
                   #AUX_rgcReceiveBuffer[13] = ' ' AND
                   #AUX_rgcReceiveBuffer[19] = ' ' AND
                   #AUX_rgcReceiveBuffer[25] = ' ' AND
                   #AUX_rgcReceiveBuffer[31] = ' ' AND
                   #AUX_rgcReceiveBuffer[37] = ' ' AND
                   #AUX_rgcReceiveBuffer[43] = ' ' AND
                   #AUX_rgcReceiveBuffer[49] = ' ' AND
                   #AUX_rgcReceiveBuffer[55] = ' ' AND
                   #AUX_rgcReceiveBuffer[61] = ' ' AND
                   #AUX_rgcReceiveBuffer[67] = ' ' AND
                   #AUX_rgcReceiveBuffer[73] = #STR_CR AND
                   #AUX_rgcReceiveBuffer[74] = #STR_LF THEN

                    //Evaluate the data of the Y telegram
                   #TMP_dTelCount :=  #AUX_tYTelegram.dTelCounter;               

                   #TMP_dTelCount += 1;

                   IF #TMP_dTelCount >= 65535 THEN
                       #TMP_dTelCount := 1;
                   END_IF; 

                   Chars_TO_Strg(Chars:=#AUX_rgcReceiveBuffer,
                                 pChars:=2,
                                 Cnt:=5,
                                 Strg=>#TMP_strValue);

                   #AUX_tYTelegram.dTelCounter := STRING_TO_DINT(#TMP_strValue); 

                   IF (#TMP_dTelCount <> #AUX_tYTelegram.dTelCounter) THEN
                       #AUX_xTelegramYMissing := 1;    
                   END_IF;

                   //Feeding pulse counter
                   Chars_TO_Strg(Chars:=#AUX_rgcReceiveBuffer,
                                 pChars:=8,
                                 Cnt:=5,
                                 Strg=>#TMP_strValue);

                   #AUX_tYTelegram.dFeedPulse_mm := STRING_TO_DINT(#TMP_strValue); 

                   //Inner limit of the observation area [mm]
                   Chars_TO_Strg(Chars:=#AUX_rgcReceiveBuffer,
                                 pChars:=14,
                                 Cnt:=5,
                                 Strg=>#TMP_strValue);

                   #AUX_tYTelegram.dInLimit_mm := STRING_TO_DINT(#TMP_strValue); 


                   //Outer limit of the observation area [mm]
                   Chars_TO_Strg(Chars:=#AUX_rgcReceiveBuffer,
                                 pChars:=20,
                                 Cnt:=5,
                                 Strg=>#TMP_strValue);

                   #AUX_tYTelegram.dOutLimit_mm := STRING_TO_DINT(#TMP_strValue); 

                   //Inner limit of the usable glass width [mm]
                   Chars_TO_Strg(Chars:=#AUX_rgcReceiveBuffer,
                                 pChars:=26,
                                 Cnt:=5,
                                 Strg=>#TMP_strValue);

                   #AUX_tYTelegram.dInLimitUsable_mm := STRING_TO_DINT(#TMP_strValue); 

                   //Outer limit of the usable glass width [mm]
                   Chars_TO_Strg(Chars:=#AUX_rgcReceiveBuffer,
                                 pChars:=32,
                                 Cnt:=5,
                                 Strg=>#TMP_strValue);

                   #AUX_tYTelegram.dOutLimitUsable_mm := STRING_TO_DINT(#TMP_strValue); 